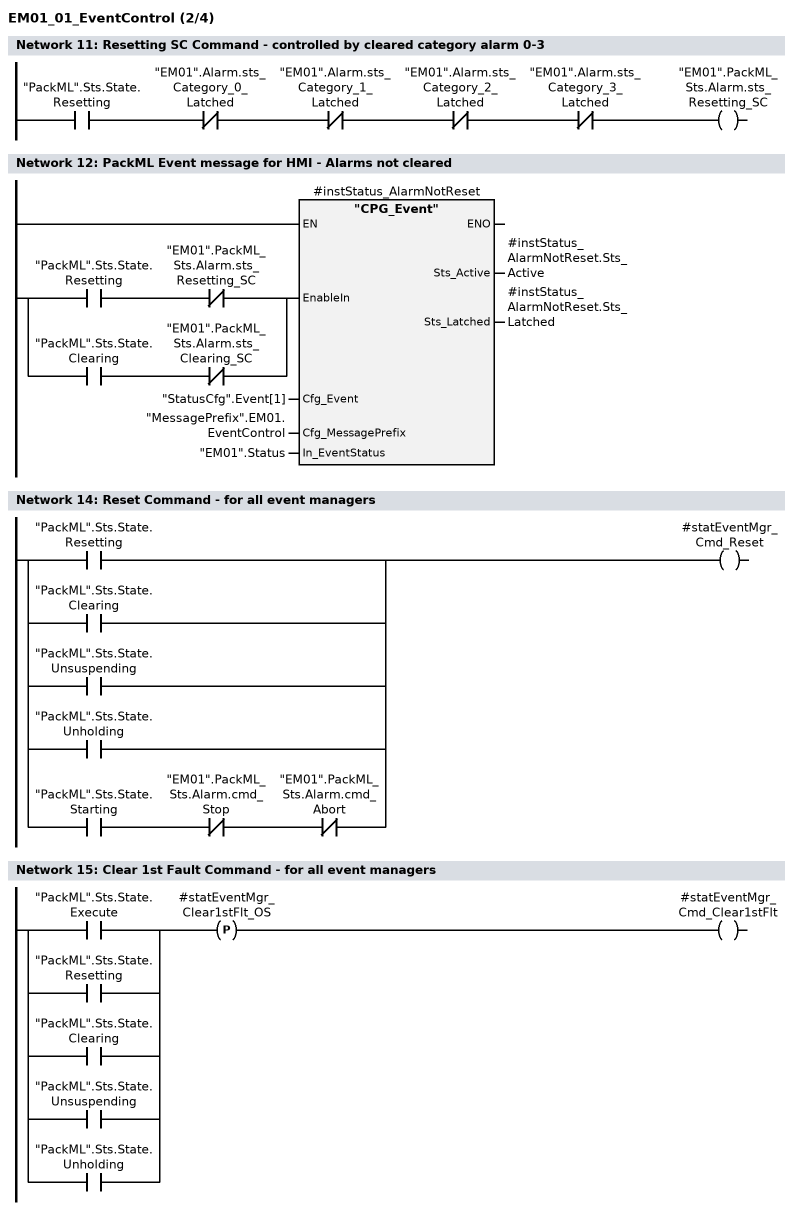
   RUNG wire#powerrail
      Contact( "PackML".Sts.State.Resetting )
      I_Contact( "EM01".Alarm.sts_Category_0_Latched )
      I_Contact( "EM01".Alarm.sts_Category_1_Latched )
      I_Contact( "EM01".Alarm.sts_Category_2_Latched )
      I_Contact( "EM01".Alarm.sts_Category_3_Latched )
      Coil( "EM01".PackML_Sts.Alarm.sts_Resetting_SC )
   END_RUNG
   // the same network as SCL:
   "EM01".PackML_Sts.Alarm.sts_Resetting_SC := "PackML".Sts.State.Resetting AND NOT "EM01".Alarm.sts_Category_0_Latched AND NOT "EM01".Alarm.sts_Category_1_Latched AND NOT "EM01".Alarm.sts_Category_2_Latched AND NOT "EM01".Alarm.sts_Category_3_Latched;
END_REGION

REGION Network 12: PackML Event message for HMI - Alarms not cleared
   RUNG wire#powerrail
      #instStatus_AlarmNotReset(EnableIn := wire#w1, Cfg_Event := "StatusCfg".Event[1], Cfg_MessagePrefix := "MessagePrefix".EM01.EventControl, In_EventStatus := "EM01".Status, Sts_Active => #instStatus_AlarmNotReset.Sts_Active, Sts_Latched => #instStatus_AlarmNotReset.Sts_Latched)
   END_RUNG
   RUNG wire#powerrail
      Contact( "PackML".Sts.State.Resetting )
      I_Contact( "EM01".PackML_Sts.Alarm.sts_Resetting_SC )
   END_RUNG wire#w1
   RUNG wire#powerrail
      Contact( "PackML".Sts.State.Clearing )
      I_Contact( "EM01".PackML_Sts.Alarm.sts_Clearing_SC )
   END_RUNG wire#w1
   // the same network as SCL:
   #instStatus_AlarmNotReset(EnableIn := ("PackML".Sts.State.Resetting AND NOT "EM01".PackML_Sts.Alarm.sts_Resetting_SC) OR ("PackML".Sts.State.Clearing AND NOT "EM01".PackML_Sts.Alarm.sts_Clearing_SC),   // "CPG_Event"
                           Cfg_Event := "StatusCfg".Event[1],
                           Cfg_MessagePrefix := "MessagePrefix".EM01.EventControl,
                           In_EventStatus := "EM01".Status,
                           Sts_Active => #instStatus_AlarmNotReset.Sts_Active,
                           Sts_Latched => #instStatus_AlarmNotReset.Sts_Latched);
END_REGION

REGION Network 13: *** EVENT CONTROL MANAGERS ***
END_REGION

REGION Network 14: Reset Command - for all event managers
   RUNG wire#powerrail
      Contact( "PackML".Sts.State.Resetting )
      wire#w1
      Coil( #statEventMgr_Cmd_Reset )
   END_RUNG
   RUNG wire#powerrail
      Contact( "PackML".Sts.State.Clearing )
   END_RUNG wire#w1
   RUNG wire#powerrail
      Contact( "PackML".Sts.State.Unsuspending )
   END_RUNG wire#w1
   RUNG wire#powerrail
      Contact( "PackML".Sts.State.Unholding )
   END_RUNG wire#w1
   RUNG wire#powerrail
      Contact( "PackML".Sts.State.Starting )
      I_Contact( "EM01".PackML_Sts.Alarm.cmd_Stop )
      I_Contact( "EM01".PackML_Sts.Alarm.cmd_Abort )
   END_RUNG wire#w1
   // the same network as SCL:
   #statEventMgr_Cmd_Reset := "PackML".Sts.State.Resetting OR "PackML".Sts.State.Clearing OR "PackML".Sts.State.Unsuspending OR "PackML".Sts.State.Unholding OR ("PackML".Sts.State.Starting AND NOT "EM01".PackML_Sts.Alarm.cmd_Stop AND NOT "EM01".PackML_Sts.Alarm.cmd_Abort);
END_REGION

REGION Network 15: Clear 1st Fault Command - for all event managers
   RUNG wire#powerrail
      Contact( "PackML".Sts.State.Execute )
      wire#w1
      P_Trig( #statEventMgr_Clear1stFlt_OS )
      Coil( #statEventMgr_Cmd_Clear1stFlt )
   END_RUNG
   RUNG wire#powerrail
      Contact( "PackML".Sts.State.Resetting )
   END_RUNG wire#w1
   RUNG wire#powerrail
      Contact( "PackML".Sts.State.Clearing )
   END_RUNG wire#w1
   RUNG wire#powerrail
      Contact( "PackML".Sts.State.Unsuspending )
   END_RUNG wire#w1
   RUNG wire#powerrail
      Contact( "PackML".Sts.State.Unholding )
   END_RUNG wire#w1
   // the same network as SCL:
   #_w1 := "PackML".Sts.State.Execute OR "PackML".Sts.State.Resetting OR "PackML".Sts.State.Clearing OR "PackML".Sts.State.Unsuspending OR "PackML".Sts.State.Unholding;
   #_w2 := #_w1 AND NOT #statEventMgr_Clear1stFlt_OS;   // rising edge
   #statEventMgr_Clear1stFlt_OS := #_w1;
   #statEventMgr_Cmd_Clear1stFlt := #_w2;
END_REGION

REGION Network 16: Call the Event Manager logic for EM alarms
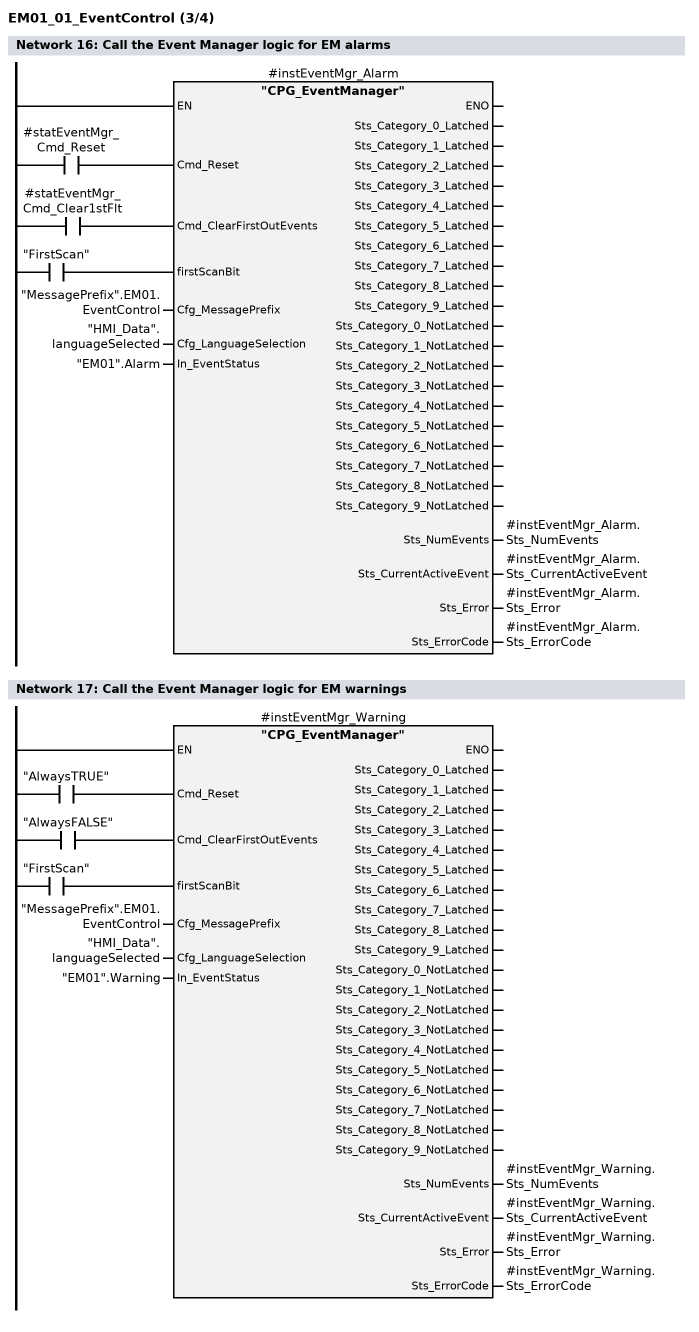
   RUNG wire#powerrail
      #instEventMgr_Alarm(Cmd_Reset := wire#w1, Cmd_ClearFirstOutEvents := wire#w2, firstScanBit := wire#w3, Cfg_MessagePrefix := "MessagePrefix".EM01.EventControl, Cfg_LanguageSelection := "HMI_Data".languageSelected, In_EventStatus := "EM01".Alarm, Sts_Category_0_Latched =>, Sts_Category_1_Latched =>, Sts_Category_2_Latched =>, Sts_Category_3_Latched =>, Sts_Category_4_Latched =>, Sts_Category_5_Latched =>, Sts_Category_6_Latched =>, Sts_Category_7_Latched =>, Sts_Category_8_Latched =>, Sts_Category_9_Latched =>, Sts_Category_0_NotLatched =>, Sts_Category_1_NotLatched =>, Sts_Category_2_NotLatched =>, Sts_Category_3_NotLatched =>, Sts_Category_4_NotLatched =>, Sts_Category_5_NotLatched =>, Sts_Category_6_NotLatched =>, Sts_Category_7_NotLatched =>, Sts_Category_8_NotLatched =>, Sts_Category_9_NotLatched =>, Sts_NumEvents => #instEventMgr_Alarm.Sts_NumEvents, Sts_CurrentActiveEvent => #instEventMgr_Alarm.Sts_CurrentActiveEvent, Sts_Error => #instEventMgr_Alarm.Sts_Error, Sts_ErrorCode => #instEventMgr_Alarm.Sts_ErrorCode)
   END_RUNG
   RUNG wire#powerrail
      Contact( #statEventMgr_Cmd_Reset )
   END_RUNG wire#w1
   RUNG wire#powerrail
      Contact( #statEventMgr_Cmd_Clear1stFlt )
   END_RUNG wire#w2
   RUNG wire#powerrail
      Contact( "FirstScan" )
   END_RUNG wire#w3
   // the same network as SCL:
   #instEventMgr_Alarm(Cmd_Reset := #statEventMgr_Cmd_Reset,   // "CPG_EventManager"
                       Cmd_ClearFirstOutEvents := #statEventMgr_Cmd_Clear1stFlt,
                       firstScanBit := "FirstScan",
                       Cfg_MessagePrefix := "MessagePrefix".EM01.EventControl,
                       Cfg_LanguageSelection := "HMI_Data".languageSelected,
                       In_EventStatus := "EM01".Alarm,
                       Sts_NumEvents => #instEventMgr_Alarm.Sts_NumEvents,
                       Sts_CurrentActiveEvent => #instEventMgr_Alarm.Sts_CurrentActiveEvent,
                       Sts_Error => #instEventMgr_Alarm.Sts_Error,
                       Sts_ErrorCode => #instEventMgr_Alarm.Sts_ErrorCode);
END_REGION

REGION Network 17: Call the Event Manager logic for EM warnings
   RUNG wire#powerrail
      #instEventMgr_Warning(Cmd_Reset := wire#w1, Cmd_ClearFirstOutEvents := wire#w2, firstScanBit := wire#w3, Cfg_MessagePrefix := "MessagePrefix".EM01.EventControl, Cfg_LanguageSelection := "HMI_Data".languageSelected, In_EventStatus := "EM01".Warning, Sts_Category_0_Latched =>, Sts_Category_1_Latched =>, Sts_Category_2_Latched =>, Sts_Category_3_Latched =>, Sts_Category_4_Latched =>, Sts_Category_5_Latched =>, Sts_Category_6_Latched =>, Sts_Category_7_Latched =>, Sts_Category_8_Latched =>, Sts_Category_9_Latched =>, Sts_Category_0_NotLatched =>, Sts_Category_1_NotLatched =>, Sts_Category_2_NotLatched =>, Sts_Category_3_NotLatched =>, Sts_Category_4_NotLatched =>, Sts_Category_5_NotLatched =>, Sts_Category_6_NotLatched =>, Sts_Category_7_NotLatched =>, Sts_Category_8_NotLatched =>, Sts_Category_9_NotLatched =>, Sts_NumEvents => #instEventMgr_Warning.Sts_NumEvents, Sts_CurrentActiveEvent => #instEventMgr_Warning.Sts_CurrentActiveEvent, Sts_Error => #instEventMgr_Warning.Sts_Error, Sts_ErrorCode => #instEventMgr_Warning.Sts_ErrorCode)
   END_RUNG
   RUNG wire#powerrail
      Contact( "AlwaysTRUE" )
   END_RUNG wire#w1
   RUNG wire#powerrail
      Contact( "AlwaysFALSE" )
   END_RUNG wire#w2
   RUNG wire#powerrail
      Contact( "FirstScan" )
   END_RUNG wire#w3
   // the same network as SCL:
   #instEventMgr_Warning(Cmd_Reset := "AlwaysTRUE",   // "CPG_EventManager"
                         Cmd_ClearFirstOutEvents := "AlwaysFALSE",
                         firstScanBit := "FirstScan",
                         Cfg_MessagePrefix := "MessagePrefix".EM01.EventControl,
                         Cfg_LanguageSelection := "HMI_Data".languageSelected,
                         In_EventStatus := "EM01".Warning,
                         Sts_NumEvents => #instEventMgr_Warning.Sts_NumEvents,
                         Sts_CurrentActiveEvent => #instEventMgr_Warning.Sts_CurrentActiveEvent,
                         Sts_Error => #instEventMgr_Warning.Sts_Error,
                         Sts_ErrorCode => #instEventMgr_Warning.Sts_ErrorCode);
END_REGION

REGION Network 18: Call the Event Manager logic for EM status
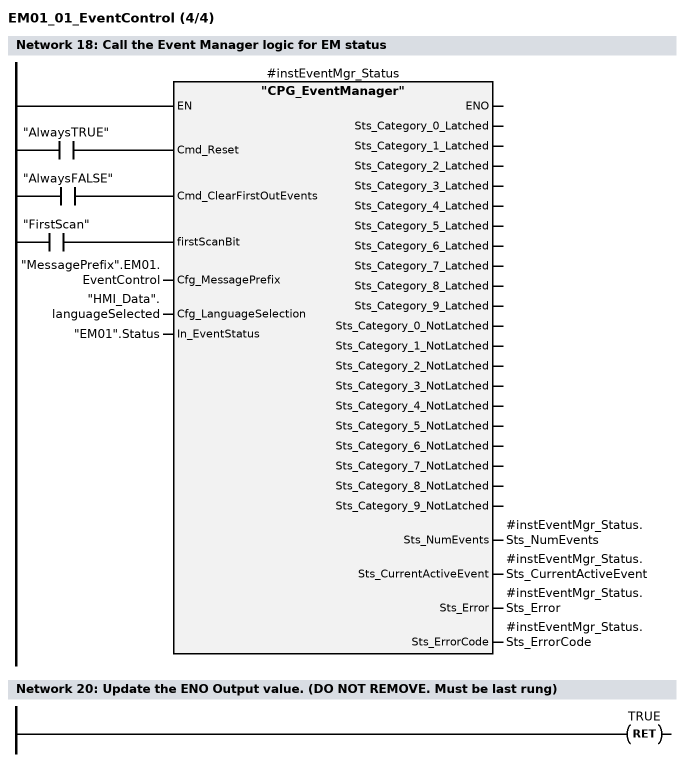
   RUNG wire#powerrail
      #instEventMgr_Status(Cmd_Reset := wire#w1, Cmd_ClearFirstOutEvents := wire#w2, firstScanBit := wire#w3, Cfg_MessagePrefix := "MessagePrefix".EM01.EventControl, Cfg_LanguageSelection := "HMI_Data".languageSelected, In_EventStatus := "EM01".Status, Sts_Category_0_Latched =>, Sts_Category_1_Latched =>, Sts_Category_2_Latched =>, Sts_Category_3_Latched =>, Sts_Category_4_Latched =>, Sts_Category_5_Latched =>, Sts_Category_6_Latched =>, Sts_Category_7_Latched =>, Sts_Category_8_Latched =>, Sts_Category_9_Latched =>, Sts_Category_0_NotLatched =>, Sts_Category_1_NotLatched =>, Sts_Category_2_NotLatched =>, Sts_Category_3_NotLatched =>, Sts_Category_4_NotLatched =>, Sts_Category_5_NotLatched =>, Sts_Category_6_NotLatched =>, Sts_Category_7_NotLatched =>, Sts_Category_8_NotLatched =>, Sts_Category_9_NotLatched =>, Sts_NumEvents => #instEventMgr_Status.Sts_NumEvents, Sts_CurrentActiveEvent => #instEventMgr_Status.Sts_CurrentActiveEvent, Sts_Error => #instEventMgr_Status.Sts_Error, Sts_ErrorCode => #instEventMgr_Status.Sts_ErrorCode)
   END_RUNG
   RUNG wire#powerrail
      Contact( "AlwaysTRUE" )
   END_RUNG wire#w1
   RUNG wire#powerrail
      Contact( "AlwaysFALSE" )
   END_RUNG wire#w2
   RUNG wire#powerrail
      Contact( "FirstScan" )
   END_RUNG wire#w3
   // the same network as SCL:
   #instEventMgr_Status(Cmd_Reset := "AlwaysTRUE",   // "CPG_EventManager"
                        Cmd_ClearFirstOutEvents := "AlwaysFALSE",
                        firstScanBit := "FirstScan",
                        Cfg_MessagePrefix := "MessagePrefix".EM01.EventControl,
                        Cfg_LanguageSelection := "HMI_Data".languageSelected,
                        In_EventStatus := "EM01".Status,
                        Sts_NumEvents => #instEventMgr_Status.Sts_NumEvents,
                        Sts_CurrentActiveEvent => #instEventMgr_Status.Sts_CurrentActiveEvent,
                        Sts_Error => #instEventMgr_Status.Sts_Error,
                        Sts_ErrorCode => #instEventMgr_Status.Sts_ErrorCode);
END_REGION

REGION Network 20: Update the ENO Output value. (DO NOT REMOVE. Must be last rung)
   RUNG wire#powerrail
      ReturnCoil( TRUE )
   END_RUNG
   // the same network as SCL:
   ENO := TRUE;
   RETURN;
END_REGION
END_FUNCTION_BLOCK

FUNCTION_BLOCK "EM01_02_PackML_ModuleSum"   // FB31662, LAD
TITLE = EM01_02_PackML_ModuleSum
{ S7_Optimized_Access := 'TRUE' }
AUTHOR : tech.team.motioncontrol@siemens.com
FAMILY : CPG
VERSION : 1.1
// Support: tech.team.motioncontrol@siemens.com
   VAR
      statDummyBool : Bool;   // dummy bool - placeholder
   END_VAR
BEGIN

REGION Network 1: EM - Reset Command
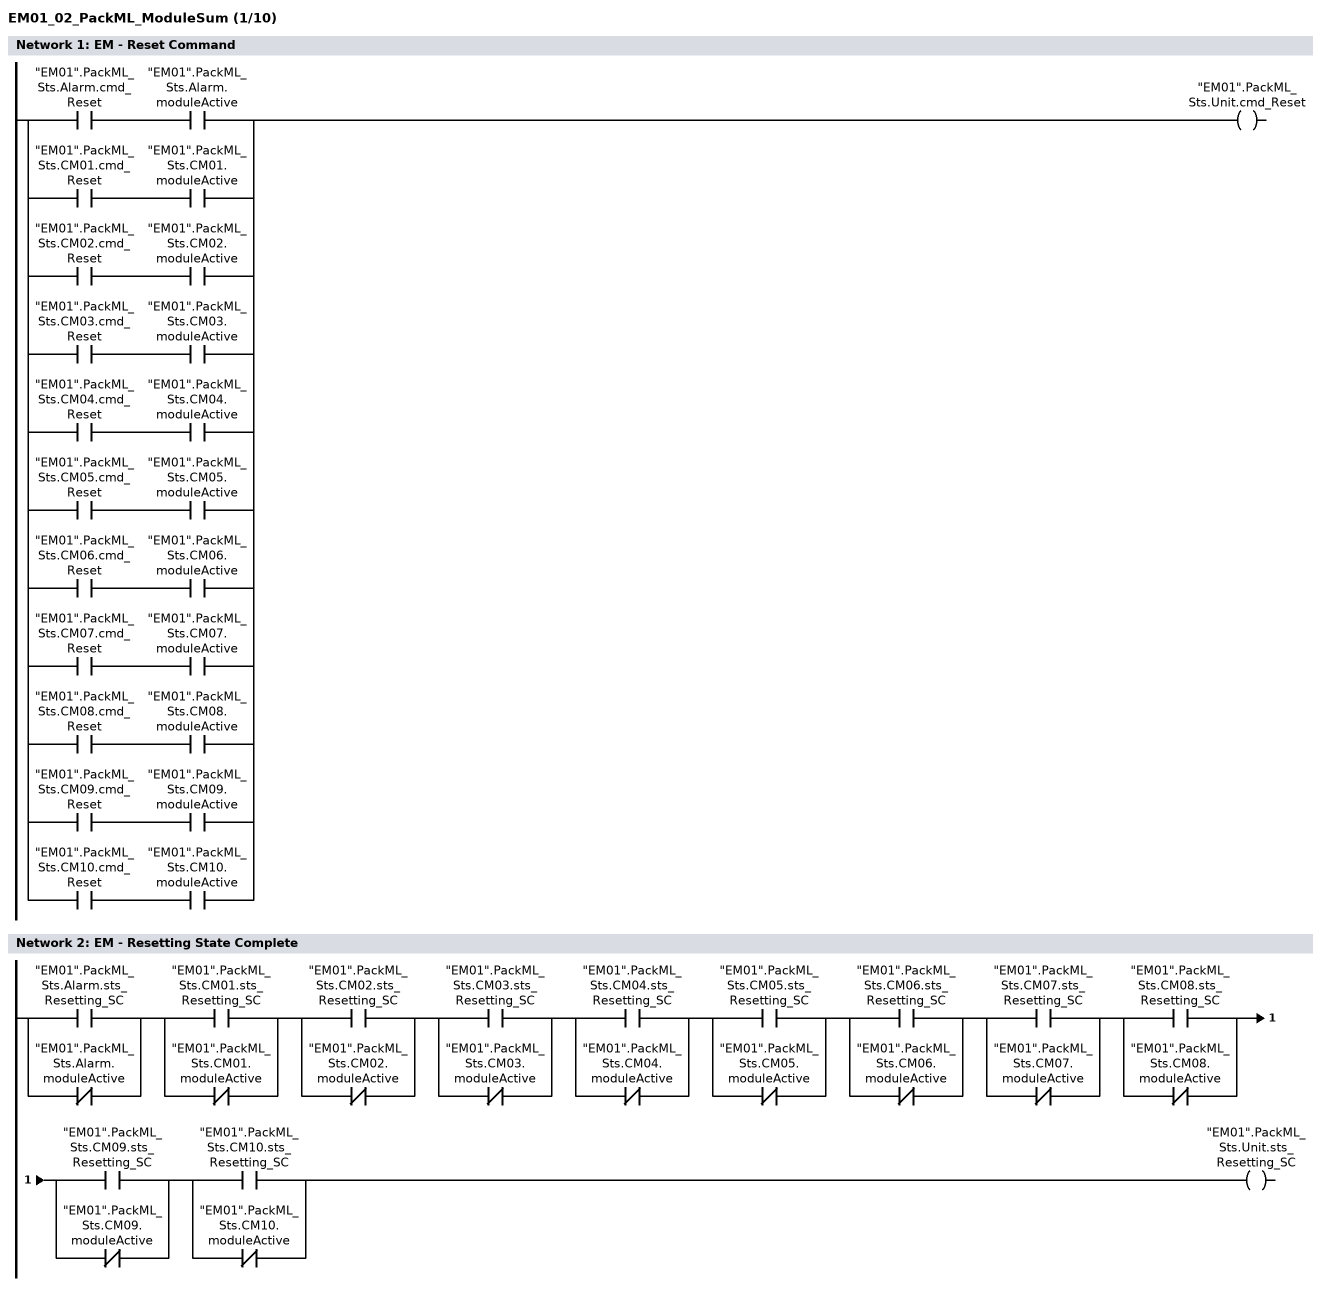
   RUNG wire#powerrail
      Contact( "EM01".PackML_Sts.Alarm.cmd_Reset )
      Contact( "EM01".PackML_Sts.Alarm.moduleActive )
      wire#w1
      Coil( "EM01".PackML_Sts.Unit.cmd_Reset )
   END_RUNG
   RUNG wire#powerrail
      Contact( "EM01".PackML_Sts.CM01.cmd_Reset )
      Contact( "EM01".PackML_Sts.CM01.moduleActive )
   END_RUNG wire#w1
   RUNG wire#powerrail
      Contact( "EM01".PackML_Sts.CM02.cmd_Reset )
      Contact( "EM01".PackML_Sts.CM02.moduleActive )
   END_RUNG wire#w1
   RUNG wire#powerrail
      Contact( "EM01".PackML_Sts.CM03.cmd_Reset )
      Contact( "EM01".PackML_Sts.CM03.moduleActive )
   END_RUNG wire#w1
   RUNG wire#powerrail
      Contact( "EM01".PackML_Sts.CM04.cmd_Reset )
      Contact( "EM01".PackML_Sts.CM04.moduleActive )
   END_RUNG wire#w1
   RUNG wire#powerrail
      Contact( "EM01".PackML_Sts.CM05.cmd_Reset )
      Contact( "EM01".PackML_Sts.CM05.moduleActive )
   END_RUNG wire#w1
   RUNG wire#powerrail
      Contact( "EM01".PackML_Sts.CM06.cmd_Reset )
      Contact( "EM01".PackML_Sts.CM06.moduleActive )
   END_RUNG wire#w1
   RUNG wire#powerrail
      Contact( "EM01".PackML_Sts.CM07.cmd_Reset )
      Contact( "EM01".PackML_Sts.CM07.moduleActive )
   END_RUNG wire#w1
   RUNG wire#powerrail
      Contact( "EM01".PackML_Sts.CM08.cmd_Reset )
      Contact( "EM01".PackML_Sts.CM08.moduleActive )
   END_RUNG wire#w1
   RUNG wire#powerrail
      Contact( "EM01".PackML_Sts.CM09.cmd_Reset )
      Contact( "EM01".PackML_Sts.CM09.moduleActive )
   END_RUNG wire#w1
   RUNG wire#powerrail
      Contact( "EM01".PackML_Sts.CM10.cmd_Reset )
      Contact( "EM01".PackML_Sts.CM10.moduleActive )
   END_RUNG wire#w1
   // the same network as SCL:
   "EM01".PackML_Sts.Unit.cmd_Reset := ("EM01".PackML_Sts.Alarm.cmd_Reset AND "EM01".PackML_Sts.Alarm.moduleActive) OR ("EM01".PackML_Sts.CM01.cmd_Reset AND "EM01".PackML_Sts.CM01.moduleActive) OR ("EM01".PackML_Sts.CM02.cmd_Reset AND "EM01".PackML_Sts.CM02.moduleActive) OR ("EM01".PackML_Sts.CM03.cmd_Reset AND "EM01".PackML_Sts.CM03.moduleActive) OR ("EM01".PackML_Sts.CM04.cmd_Reset AND "EM01".PackML_Sts.CM04.moduleActive) OR ("EM01".PackML_Sts.CM05.cmd_Reset AND "EM01".PackML_Sts.CM05.moduleActive) OR ("EM01".PackML_Sts.CM06.cmd_Reset AND "EM01".PackML_Sts.CM06.moduleActive) OR ("EM01".PackML_Sts.CM07.cmd_Reset AND "EM01".PackML_Sts.CM07.moduleActive) OR ("EM01".PackML_Sts.CM08.cmd_Reset AND "EM01".PackML_Sts.CM08.moduleActive) OR ("EM01".PackML_Sts.CM09.cmd_Reset AND "EM01".PackML_Sts.CM09.moduleActive) OR ("EM01".PackML_Sts.CM10.cmd_Reset AND "EM01".PackML_Sts.CM10.moduleActive);
END_REGION

REGION Network 2: EM - Resetting State Complete
   RUNG wire#powerrail
      Contact( "EM01".PackML_Sts.Alarm.sts_Resetting_SC )
      wire#w1
      Contact( "EM01".PackML_Sts.CM01.sts_Resetting_SC )
      wire#w2
      Contact( "EM01".PackML_Sts.CM02.sts_Resetting_SC )
      wire#w3
      Contact( "EM01".PackML_Sts.CM03.sts_Resetting_SC )
      wire#w4
      Contact( "EM01".PackML_Sts.CM04.sts_Resetting_SC )
      wire#w5
      Contact( "EM01".PackML_Sts.CM05.sts_Resetting_SC )
      wire#w6
      Contact( "EM01".PackML_Sts.CM06.sts_Resetting_SC )
      wire#w7
      Contact( "EM01".PackML_Sts.CM07.sts_Resetting_SC )
      wire#w8
      Contact( "EM01".PackML_Sts.CM08.sts_Resetting_SC )
      wire#w9
      Contact( "EM01".PackML_Sts.CM09.sts_Resetting_SC )
      wire#w10
      Contact( "EM01".PackML_Sts.CM10.sts_Resetting_SC )
      wire#w11
      Coil( "EM01".PackML_Sts.Unit.sts_Resetting_SC )
   END_RUNG
   RUNG wire#powerrail
      I_Contact( "EM01".PackML_Sts.Alarm.moduleActive )
   END_RUNG wire#w1
   RUNG wire#w1
      I_Contact( "EM01".PackML_Sts.CM01.moduleActive )
   END_RUNG wire#w2
   RUNG wire#w2
      I_Contact( "EM01".PackML_Sts.CM02.moduleActive )
   END_RUNG wire#w3
   RUNG wire#w3
      I_Contact( "EM01".PackML_Sts.CM03.moduleActive )
   END_RUNG wire#w4
   RUNG wire#w4
      I_Contact( "EM01".PackML_Sts.CM04.moduleActive )
   END_RUNG wire#w5
   RUNG wire#w5
      I_Contact( "EM01".PackML_Sts.CM05.moduleActive )
   END_RUNG wire#w6
   RUNG wire#w6
      I_Contact( "EM01".PackML_Sts.CM06.moduleActive )
   END_RUNG wire#w7
   RUNG wire#w7
      I_Contact( "EM01".PackML_Sts.CM07.moduleActive )
   END_RUNG wire#w8
   RUNG wire#w8
      I_Contact( "EM01".PackML_Sts.CM08.moduleActive )
   END_RUNG wire#w9
   RUNG wire#w9
      I_Contact( "EM01".PackML_Sts.CM09.moduleActive )
   END_RUNG wire#w10
   RUNG wire#w10
      I_Contact( "EM01".PackML_Sts.CM10.moduleActive )
   END_RUNG wire#w11
   // the same network as SCL:
   "EM01".PackML_Sts.Unit.sts_Resetting_SC := ("EM01".PackML_Sts.Alarm.sts_Resetting_SC OR NOT "EM01".PackML_Sts.Alarm.moduleActive) AND ("EM01".PackML_Sts.CM01.sts_Resetting_SC OR NOT "EM01".PackML_Sts.CM01.moduleActive) AND ("EM01".PackML_Sts.CM02.sts_Resetting_SC OR NOT "EM01".PackML_Sts.CM02.moduleActive) AND ("EM01".PackML_Sts.CM03.sts_Resetting_SC OR NOT "EM01".PackML_Sts.CM03.moduleActive) AND ("EM01".PackML_Sts.CM04.sts_Resetting_SC OR NOT "EM01".PackML_Sts.CM04.moduleActive) AND ("EM01".PackML_Sts.CM05.sts_Resetting_SC OR NOT "EM01".PackML_Sts.CM05.moduleActive) AND ("EM01".PackML_Sts.CM06.sts_Resetting_SC OR NOT "EM01".PackML_Sts.CM06.moduleActive) AND ("EM01".PackML_Sts.CM07.sts_Resetting_SC OR NOT "EM01".PackML_Sts.CM07.moduleActive) AND ("EM01".PackML_Sts.CM08.sts_Resetting_SC OR NOT "EM01".PackML_Sts.CM08.moduleActive) AND ("EM01".PackML_Sts.CM09.sts_Resetting_SC OR NOT "EM01".PackML_Sts.CM09.moduleActive) AND ("EM01".PackML_Sts.CM10.sts_Resetting_SC OR NOT "EM01".PackML_Sts.CM10.moduleActive);
END_REGION

REGION Network 3: EM - Start Command
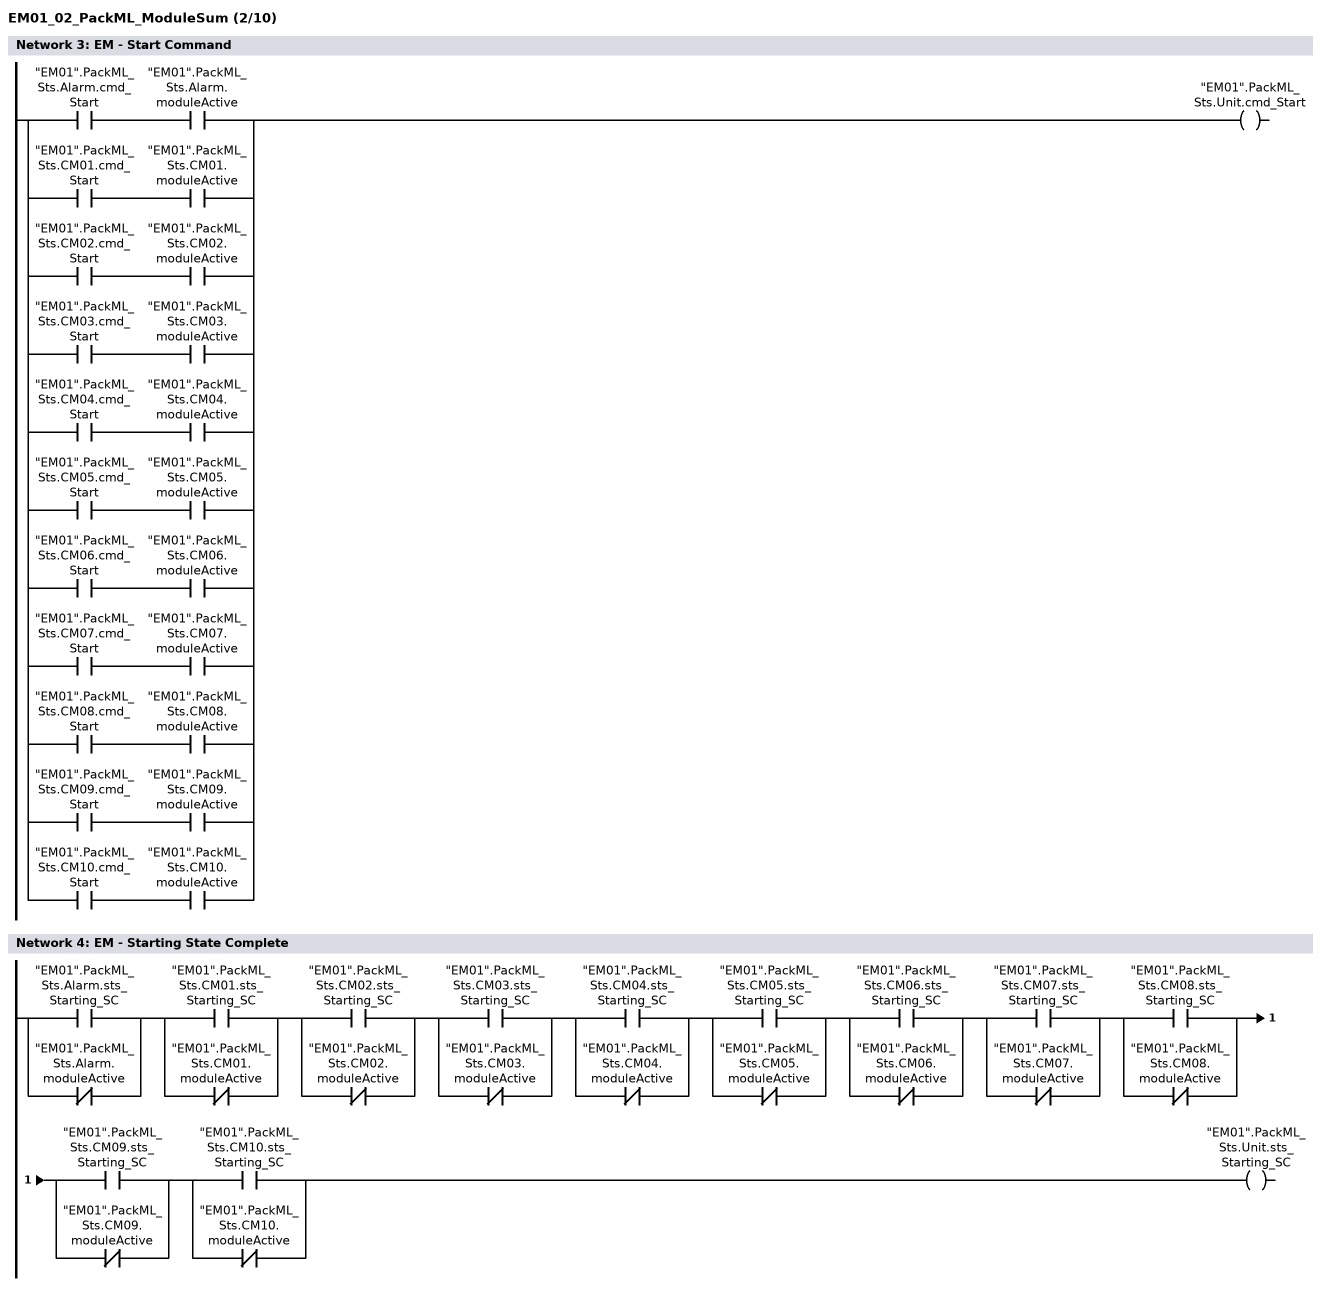
   RUNG wire#powerrail
      Contact( "EM01".PackML_Sts.Alarm.cmd_Start )
      Contact( "EM01".PackML_Sts.Alarm.moduleActive )
      wire#w1
      Coil( "EM01".PackML_Sts.Unit.cmd_Start )
   END_RUNG
   RUNG wire#powerrail
      Contact( "EM01".PackML_Sts.CM01.cmd_Start )
      Contact( "EM01".PackML_Sts.CM01.moduleActive )
   END_RUNG wire#w1
   RUNG wire#powerrail
      Contact( "EM01".PackML_Sts.CM02.cmd_Start )
      Contact( "EM01".PackML_Sts.CM02.moduleActive )
   END_RUNG wire#w1
   RUNG wire#powerrail
      Contact( "EM01".PackML_Sts.CM03.cmd_Start )
      Contact( "EM01".PackML_Sts.CM03.moduleActive )
   END_RUNG wire#w1
   RUNG wire#powerrail
      Contact( "EM01".PackML_Sts.CM04.cmd_Start )
      Contact( "EM01".PackML_Sts.CM04.moduleActive )
   END_RUNG wire#w1
   RUNG wire#powerrail
      Contact( "EM01".PackML_Sts.CM05.cmd_Start )
      Contact( "EM01".PackML_Sts.CM05.moduleActive )
   END_RUNG wire#w1
   RUNG wire#powerrail
      Contact( "EM01".PackML_Sts.CM06.cmd_Start )
      Contact( "EM01".PackML_Sts.CM06.moduleActive )
   END_RUNG wire#w1
   RUNG wire#powerrail
      Contact( "EM01".PackML_Sts.CM07.cmd_Start )
      Contact( "EM01".PackML_Sts.CM07.moduleActive )
   END_RUNG wire#w1
   RUNG wire#powerrail
      Contact( "EM01".PackML_Sts.CM08.cmd_Start )
      Contact( "EM01".PackML_Sts.CM08.moduleActive )
   END_RUNG wire#w1
   RUNG wire#powerrail
      Contact( "EM01".PackML_Sts.CM09.cmd_Start )
      Contact( "EM01".PackML_Sts.CM09.moduleActive )
   END_RUNG wire#w1
   RUNG wire#powerrail
      Contact( "EM01".PackML_Sts.CM10.cmd_Start )
      Contact( "EM01".PackML_Sts.CM10.moduleActive )
   END_RUNG wire#w1
   // the same network as SCL:
   "EM01".PackML_Sts.Unit.cmd_Start := ("EM01".PackML_Sts.Alarm.cmd_Start AND "EM01".PackML_Sts.Alarm.moduleActive) OR ("EM01".PackML_Sts.CM01.cmd_Start AND "EM01".PackML_Sts.CM01.moduleActive) OR ("EM01".PackML_Sts.CM02.cmd_Start AND "EM01".PackML_Sts.CM02.moduleActive) OR ("EM01".PackML_Sts.CM03.cmd_Start AND "EM01".PackML_Sts.CM03.moduleActive) OR ("EM01".PackML_Sts.CM04.cmd_Start AND "EM01".PackML_Sts.CM04.moduleActive) OR ("EM01".PackML_Sts.CM05.cmd_Start AND "EM01".PackML_Sts.CM05.moduleActive) OR ("EM01".PackML_Sts.CM06.cmd_Start AND "EM01".PackML_Sts.CM06.moduleActive) OR ("EM01".PackML_Sts.CM07.cmd_Start AND "EM01".PackML_Sts.CM07.moduleActive) OR ("EM01".PackML_Sts.CM08.cmd_Start AND "EM01".PackML_Sts.CM08.moduleActive) OR ("EM01".PackML_Sts.CM09.cmd_Start AND "EM01".PackML_Sts.CM09.moduleActive) OR ("EM01".PackML_Sts.CM10.cmd_Start AND "EM01".PackML_Sts.CM10.moduleActive);
END_REGION

REGION Network 4: EM - Starting State Complete
   RUNG wire#powerrail
      Contact( "EM01".PackML_Sts.Alarm.sts_Starting_SC )
      wire#w1
      Contact( "EM01".PackML_Sts.CM01.sts_Starting_SC )
      wire#w2
      Contact( "EM01".PackML_Sts.CM02.sts_Starting_SC )
      wire#w3
      Contact( "EM01".PackML_Sts.CM03.sts_Starting_SC )
      wire#w4
      Contact( "EM01".PackML_Sts.CM04.sts_Starting_SC )
      wire#w5
      Contact( "EM01".PackML_Sts.CM05.sts_Starting_SC )
      wire#w6
      Contact( "EM01".PackML_Sts.CM06.sts_Starting_SC )
      wire#w7
      Contact( "EM01".PackML_Sts.CM07.sts_Starting_SC )
      wire#w8
      Contact( "EM01".PackML_Sts.CM08.sts_Starting_SC )
      wire#w9
      Contact( "EM01".PackML_Sts.CM09.sts_Starting_SC )
      wire#w10
      Contact( "EM01".PackML_Sts.CM10.sts_Starting_SC )
      wire#w11
      Coil( "EM01".PackML_Sts.Unit.sts_Starting_SC )
   END_RUNG
   RUNG wire#powerrail
      I_Contact( "EM01".PackML_Sts.Alarm.moduleActive )
   END_RUNG wire#w1
   RUNG wire#w1
      I_Contact( "EM01".PackML_Sts.CM01.moduleActive )
   END_RUNG wire#w2
   RUNG wire#w2
      I_Contact( "EM01".PackML_Sts.CM02.moduleActive )
   END_RUNG wire#w3
   RUNG wire#w3
      I_Contact( "EM01".PackML_Sts.CM03.moduleActive )
   END_RUNG wire#w4
   RUNG wire#w4
      I_Contact( "EM01".PackML_Sts.CM04.moduleActive )
   END_RUNG wire#w5
   RUNG wire#w5
      I_Contact( "EM01".PackML_Sts.CM05.moduleActive )
   END_RUNG wire#w6
   RUNG wire#w6
      I_Contact( "EM01".PackML_Sts.CM06.moduleActive )
   END_RUNG wire#w7
   RUNG wire#w7
      I_Contact( "EM01".PackML_Sts.CM07.moduleActive )
   END_RUNG wire#w8
   RUNG wire#w8
      I_Contact( "EM01".PackML_Sts.CM08.moduleActive )
   END_RUNG wire#w9
   RUNG wire#w9
      I_Contact( "EM01".PackML_Sts.CM09.moduleActive )
   END_RUNG wire#w10
   RUNG wire#w10
      I_Contact( "EM01".PackML_Sts.CM10.moduleActive )
   END_RUNG wire#w11
   // the same network as SCL:
   "EM01".PackML_Sts.Unit.sts_Starting_SC := ("EM01".PackML_Sts.Alarm.sts_Starting_SC OR NOT "EM01".PackML_Sts.Alarm.moduleActive) AND ("EM01".PackML_Sts.CM01.sts_Starting_SC OR NOT "EM01".PackML_Sts.CM01.moduleActive) AND ("EM01".PackML_Sts.CM02.sts_Starting_SC OR NOT "EM01".PackML_Sts.CM02.moduleActive) AND ("EM01".PackML_Sts.CM03.sts_Starting_SC OR NOT "EM01".PackML_Sts.CM03.moduleActive) AND ("EM01".PackML_Sts.CM04.sts_Starting_SC OR NOT "EM01".PackML_Sts.CM04.moduleActive) AND ("EM01".PackML_Sts.CM05.sts_Starting_SC OR NOT "EM01".PackML_Sts.CM05.moduleActive) AND ("EM01".PackML_Sts.CM06.sts_Starting_SC OR NOT "EM01".PackML_Sts.CM06.moduleActive) AND ("EM01".PackML_Sts.CM07.sts_Starting_SC OR NOT "EM01".PackML_Sts.CM07.moduleActive) AND ("EM01".PackML_Sts.CM08.sts_Starting_SC OR NOT "EM01".PackML_Sts.CM08.moduleActive) AND ("EM01".PackML_Sts.CM09.sts_Starting_SC OR NOT "EM01".PackML_Sts.CM09.moduleActive) AND ("EM01".PackML_Sts.CM10.sts_Starting_SC OR NOT "EM01".PackML_Sts.CM10.moduleActive);
END_REGION

REGION Network 5: EM - Stop Command